   "Carrier_44_SpareOutput(5_5)" AT %I2568.5 : Bool;   // SPARE OUTPUT
   "Carrier_44_SpareOutput(5_6)" AT %I2568.6 : Bool;   // SPARE OUTPUT
   "Carrier_44_SpareOutput(5_7)" AT %I2568.7 : Bool;   // SPARE OUTPUT
   "Carrier_44_ActualSpeed" AT %IW2570 : Word;   // ACTUAL SPEED
   "Carrier_44_CarrierDriveAlarm" AT %IW2572 : Word;   // CARRIER DRIVE ALARM
   "Carrier_44_CarrierDriveWarning" AT %IW2574 : Word;   // CARRIER DRIVE WARNING
   "Carrier_45_Status" AT %IW2600 : Word;   // CARRIER STATUS WORD
   "Carrier_45_Status.0" AT %I2600.0 : Bool;   // HEARTBEAT
   "Carrier_45_Status.1" AT %I2600.1 : Bool;   // MANUAL
   "Carrier_45_Status.2" AT %I2600.2 : Bool;   // IN_AUTO
   "Carrier_45_Status.3" AT %I2600.3 : Bool;   // POSITIONING_COMPLETE
   "Carrier_45_Status.4" AT %I2600.4 : Bool;   // PRODUCTION HOLD
   "Carrier_45_Status.5" AT %I2600.5 : Bool;   // CARRIER MOVING FORWARD
   "Carrier_45_Status.6" AT %I2600.6 : Bool;   // CARRIER MOVING REVERSE
   "Carrier_45_Status.7" AT %I2600.7 : Bool;   // CARRIER FAULT
   "Carrier_45_Status.8" AT %I2601.0 : Bool;   // CRASH DETECT TRIPPED
   "Carrier_45_Status.9" AT %I2601.1 : Bool;
   "Carrier_45_Status.10" AT %I2601.2 : Bool;
   "Carrier_45_Status.11" AT %I2601.3 : Bool;
   "Carrier_45_Status.12" AT %I2601.4 : Bool;
   "Carrier_45_Status.13" AT %I2601.5 : Bool;
   "Carrier_45_Status.14" AT %I2601.6 : Bool;
   "Carrier_45_Status.15" AT %I2601.7 : Bool;
   "Carrier_45_SDCFaultCode" AT %IW2602 : Word;   // SDC FAULT CODE
   "Carrier_45_CarrierPosition" AT %ID2604 : DWord;   // CARRIER POSITION
   "Carrier_45_CarrierNumber" AT %IW2608 : Word;   // CARRIER NUMBER
   "Carrier_45_G120DControlWord" AT %IW2610 : Word;   // G120D_STW1_CONTROL
   "Carrier_45_G120DControlWord.0" AT %I2610.0 : Bool;   // Bit_00_ON
   "Carrier_45_G120DControlWord.1" AT %I2610.1 : Bool;   // Bit_01_AUS2_INH
   "Carrier_45_G120DControlWord.2" AT %I2610.2 : Bool;   // Bit_02_AUS3_STOP
   "Carrier_45_G120DControlWord.3" AT %I2610.3 : Bool;   // Bit_03_EN
   "Carrier_45_G120DControlWord.4" AT %I2610.4 : Bool;   // Bit_04_EN_RAMP
   "Carrier_45_G120DControlWord.5" AT %I2610.5 : Bool;   // Bit_05_START_RAMP
   "Carrier_45_G120DControlWord.6" AT %I2610.6 : Bool;   // Bit_06_SETPOINT
   "Carrier_45_G120DControlWord.7" AT %I2610.7 : Bool;   // Bit_07_RESET
   "Carrier_45_G120DControlWord.8" AT %I2611.0 : Bool;   // Bit_08_JOG_R
   "Carrier_45_G120DControlWord.9" AT %I2611.1 : Bool;   // Bit_09_JOG_L
   "Carrier_45_G120DControlWord.10" AT %I2611.2 : Bool;   // Bit_10_CONTR_PLC
   "Carrier_45_G120DControlWord.11" AT %I2611.3 : Bool;   // Bit_11_REVERSE
   "Carrier_45_G120DControlWord.12" AT %I2611.4 : Bool;   // Bit_12_BRAKE_RELEASE
   "Carrier_45_G120DControlWord.13" AT %I2611.5 : Bool;   // Bit_13_DDS
   "Carrier_45_G120DControlWord.14" AT %I2611.6 : Bool;   // Bit_14_DO0
   "Carrier_45_G120DControlWord.15" AT %I2611.7 : Bool;   // Bit_15_DO1
   "Carrier_45_G120DStatusWord" AT %IW2612 : Word;   // G120D_ZSW1_STATUS
   "Carrier_45_G120DStatusWord.0" AT %I2612.0 : Bool;   // Bit_00_READY_RUN
   "Carrier_45_G120DStatusWord.1" AT %I2612.1 : Bool;   // Bit_01_READY_ON
   "Carrier_45_G120DStatusWord.2" AT %I2612.2 : Bool;   // Bit_02_ENABLE
   "Carrier_45_G120DStatusWord.3" AT %I2612.3 : Bool;   // Bit_03_FAULT
   "Carrier_45_G120DStatusWord.4" AT %I2612.4 : Bool;   // Bit_04_OFF2
   "Carrier_45_G120DStatusWord.5" AT %I2612.5 : Bool;   // Bit_05_OFF3
   "Carrier_45_G120DStatusWord.6" AT %I2612.6 : Bool;   // Bit_06_LOCK_OUT
   "Carrier_45_G120DStatusWord.7" AT %I2612.7 : Bool;   // Bit_07_WARN
   "Carrier_45_G120DStatusWord.8" AT %I2613.0 : Bool;   // Bit_08_NO_DEVIATION
   "Carrier_45_G120DStatusWord.9" AT %I2613.1 : Bool;   // Bit_09_CONTR_PLC
   "Carrier_45_G120DStatusWord.10" AT %I2613.2 : Bool;   // Bit_10_F_MAX
   "Carrier_45_G120DStatusWord.11" AT %I2613.3 : Bool;   // Bit_11_LIMIT_REACHED
   "Carrier_45_G120DStatusWord.12" AT %I2613.4 : Bool;   // Bit_12_BRAKE_OPEN
   "Carrier_45_G120DStatusWord.13" AT %I2613.5 : Bool;   // Bit_13_NO_OVERTEMP
   "Carrier_45_G120DStatusWord.14" AT %I2613.6 : Bool;   // Bit_14_CW_CCW
   "Carrier_45_G120DStatusWord.15" AT %I2613.7 : Bool;   // Bit_15_OVERL
   "Carrier_45_Slot2_Input" AT %IW2614 : Word;   // SLOT 2 INPUT WORD
   "Carrier_45_CrashDetectSW" AT %I2614.0 : Bool;   // CRASH DETECT SW
   "Carrier_45_SpareSafetyInput(2_1)" AT %I2614.1 : Bool;   // SPARE SAFETY INPUT
   "Carrier_45_SpareSafetyInput(2_2)" AT %I2614.2 : Bool;   // SPARE SAFETY INPUT
   "Carrier_45_SpareSafetyInput(2_3)" AT %I2614.3 : Bool;   // SPARE SAFETY INPUT
   "Carrier_45_SpareSafetyInput(2_4)" AT %I2614.4 : Bool;   // SPARE SAFETY INPUT
   "Carrier_45_SpareSafetyInput(2_5)" AT %I2614.5 : Bool;   // SPARE SAFETY INPUT
   "Carrier_45_SpareSafetyInput(2_6)" AT %I2614.6 : Bool;   // SPARE SAFETY INPUT
   "Carrier_45_SpareSafetyInput(2_7)" AT %I2614.7 : Bool;   // SPARE SAFETY INPUT
   "Carrier_45_Slot3_SafetyOutput" AT %IW2615 : Word;   // SLOT 3 SAFETY OUTPUT WORD
   "Carrier_45_Crash_Detect_OK" AT %I2615.0 : Bool;   // CARRIER CRASH DETECT
   "Carrier_45_SpareSafetyOutput(3_1)" AT %I2615.1 : Bool;   // SPARE SAFETY OUTPUT
   "Carrier_45_SpareSafetyOutput(3_2)" AT %I2615.2 : Bool;   // SPARE SAFETY OUTPUT
   "Carrier_45_SpareSafetyOutput(3_3)" AT %I2615.3 : Bool;   // SPARE SAFETY OUTPUT
   "Carrier_45_SpareSafetyOutput(3_4)" AT %I2615.4 : Bool;   // SPARE SAFETY OUTPUT
   "Carrier_45_SpareSafetyOutput(3_5)" AT %I2615.5 : Bool;   // SPARE SAFETY OUTPUT
   "Carrier_45_SpareSafetyOutput(3_6)" AT %I2615.6 : Bool;   // SPARE SAFETY OUTPUT
   "Carrier_45_SpareSafetyOutput(3_7)" AT %I2615.7 : Bool;   // SPARE SAFETY OUTPUT
   "Carrier_45_Slot4_Input" AT %IW2616 : Word;   // SLOT 4 INPUT WORD
   "Carrier_45_480VPowerOn_MDCB1" AT %I2616.0 : Bool;   // 480 VAC POWER ON MDCB 1
   "Carrier_45_SpareInput(4_1)" AT %I2616.1 : Bool;   // SPARE INPUT
   "Carrier_45_SpareInput(4_2)" AT %I2616.2 : Bool;   // SPARE INPUT
   "Carrier_45_SitopSelectStatus" AT %I2616.3 : Bool;   // SITOP SELECT STATUS
   "Carrier_45_DCsupplyOnPSCB2" AT %I2616.4 : Bool;   // DC SUPPLY ON PSCB 2
   "Carrier_45_SpareInput(4_5)" AT %I2616.5 : Bool;   // SPARE INPUT
   "Carrier_45_SpareInput(4_6)" AT %I2616.6 : Bool;   // SPARE INPUT
   "Carrier_45_SpareInput(4_7)" AT %I2616.7 : Bool;   // SPARE INPUT
   "Carrier_45_PB1_ProdHoldLH" AT %I2617.0 : Bool;   // PB 1 PRODUCTION HOLD LH
   "Carrier_45_PB2_ResetLH" AT %I2617.1 : Bool;   // PB 2 RESET LH
   "Carrier_45_PB3_ProdHoldRH" AT %I2617.2 : Bool;   // PB 3 PRODUCTION HOLD RH
   "Carrier_45_PB4_ResetRH" AT %I2617.3 : Bool;   // PB 4 RESET RH
   "Carrier_45_SpareInput(4_14)" AT %I2617.4 : Bool;   // SPARE INPUT
   "Carrier_45_SpareInput(4_15)" AT %I2617.5 : Bool;   // SPARE INPUT
   "Carrier_45_SpareInput(4_16)" AT %I2617.6 : Bool;   // SPARE INPUT
   "Carrier_45_SpareInput(4_17)" AT %I2617.7 : Bool;   // SPARE INPUT
   "Carrier_45_Slot5_Output" AT %IW2618 : Word;   // SLOT 5 OUTPUT WORD
   "Carrier_45_IRD400_HMI_24VDC_ENABLE" AT %I2618.0 : Bool;   // IRD 400 PANEL HMI 24V DC POWER
   "Carrier_45_FaultLight_LH" AT %I2618.1 : Bool;   // FAULT LIGHT LH
   "Carrier_45_RunLight_LH" AT %I2618.2 : Bool;   // RUN LIGHT LH
   "Carrier_45_FaultLight_RH" AT %I2618.3 : Bool;   // FAULT LIGHT RH
   "Carrier_45_RunLight_RH" AT %I2618.4 : Bool;   // RUN LIGHT RH
   "Carrier_45_SpareOutput(5_5)" AT %I2618.5 : Bool;   // SPARE OUTPUT
   "Carrier_45_SpareOutput(5_6)" AT %I2618.6 : Bool;   // SPARE OUTPUT
   "Carrier_45_SpareOutput(5_7)" AT %I2618.7 : Bool;   // SPARE OUTPUT
   "Carrier_45_ActualSpeed" AT %IW2620 : Word;   // ACTUAL SPEED
   "Carrier_45_CarrierDriveAlarm" AT %IW2622 : Word;   // CARRIER DRIVE ALARM
   "Carrier_45_CarrierDriveWarning" AT %IW2624 : Word;   // CARRIER DRIVE WARNING
   "Carrier_46_Status" AT %IW2650 : Word;   // CARRIER STATUS WORD
   "Carrier_46_Status.0" AT %I2650.0 : Bool;   // HEARTBEAT
   "Carrier_46_Status.1" AT %I2650.1 : Bool;   // MANUAL
   "Carrier_46_Status.2" AT %I2650.2 : Bool;   // IN_AUTO
   "Carrier_46_Status.3" AT %I2650.3 : Bool;   // POSITIONING_COMPLETE
   "Carrier_46_Status.4" AT %I2650.4 : Bool;   // PRODUCTION HOLD
   "Carrier_46_Status.5" AT %I2650.5 : Bool;   // CARRIER MOVING FORWARD
   "Carrier_46_Status.6" AT %I2650.6 : Bool;   // CARRIER MOVING REVERSE
   "Carrier_46_Status.7" AT %I2650.7 : Bool;   // CARRIER FAULT
   "Carrier_46_Status.8" AT %I2651.0 : Bool;   // CRASH DETECT TRIPPED
   "Carrier_46_Status.9" AT %I2651.1 : Bool;
   "Carrier_46_Status.10" AT %I2651.2 : Bool;
   "Carrier_46_Status.11" AT %I2651.3 : Bool;
   "Carrier_46_Status.12" AT %I2651.4 : Bool;
   "Carrier_46_Status.13" AT %I2651.5 : Bool;
   "Carrier_46_Status.14" AT %I2651.6 : Bool;
   "Carrier_46_Status.15" AT %I2651.7 : Bool;
   "Carrier_46_SDCFaultCode" AT %IW2652 : Word;   // SDC FAULT CODE
   "Carrier_46_CarrierPosition" AT %ID2654 : DWord;   // CARRIER POSITION
   "Carrier_46_CarrierNumber" AT %IW2658 : Word;   // CARRIER NUMBER
   "Carrier_46_G120DControlWord" AT %IW2660 : Word;   // G120D_STW1_CONTROL
   "Carrier_46_G120DControlWord.0" AT %I2660.0 : Bool;   // Bit_00_ON
   "Carrier_46_G120DControlWord.1" AT %I2660.1 : Bool;   // Bit_01_AUS2_INH
   "Carrier_46_G120DControlWord.2" AT %I2660.2 : Bool;   // Bit_02_AUS3_STOP
   "Carrier_46_G120DControlWord.3" AT %I2660.3 : Bool;   // Bit_03_EN
   "Carrier_46_G120DControlWord.4" AT %I2660.4 : Bool;   // Bit_04_EN_RAMP
   "Carrier_46_G120DControlWord.5" AT %I2660.5 : Bool;   // Bit_05_START_RAMP
   "Carrier_46_G120DControlWord.6" AT %I2660.6 : Bool;   // Bit_06_SETPOINT
   "Carrier_46_G120DControlWord.7" AT %I2660.7 : Bool;   // Bit_07_RESET
   "Carrier_46_G120DControlWord.8" AT %I2661.0 : Bool;   // Bit_08_JOG_R
   "Carrier_46_G120DControlWord.9" AT %I2661.1 : Bool;   // Bit_09_JOG_L
   "Carrier_46_G120DControlWord.10" AT %I2661.2 : Bool;   // Bit_10_CONTR_PLC
   "Carrier_46_G120DControlWord.11" AT %I2661.3 : Bool;   // Bit_11_REVERSE
   "Carrier_46_G120DControlWord.12" AT %I2661.4 : Bool;   // Bit_12_BRAKE_RELEASE
   "Carrier_46_G120DControlWord.13" AT %I2661.5 : Bool;   // Bit_13_DDS
   "Carrier_46_G120DControlWord.14" AT %I2661.6 : Bool;   // Bit_14_DO0
   "Carrier_46_G120DControlWord.15" AT %I2661.7 : Bool;   // Bit_15_DO1
   "Carrier_46_G120DStatusWord" AT %IW2662 : Word;   // G120D_ZSW1_STATUS
   "Carrier_46_G120DStatusWord.0" AT %I2662.0 : Bool;   // Bit_00_READY_RUN
   "Carrier_46_G120DStatusWord.1" AT %I2662.1 : Bool;   // Bit_01_READY_ON
   "Carrier_46_G120DStatusWord.2" AT %I2662.2 : Bool;   // Bit_02_ENABLE
   "Carrier_46_G120DStatusWord.3" AT %I2662.3 : Bool;   // Bit_03_FAULT
   "Carrier_46_G120DStatusWord.4" AT %I2662.4 : Bool;   // Bit_04_OFF2
   "Carrier_46_G120DStatusWord.5" AT %I2662.5 : Bool;   // Bit_05_OFF3
   "Carrier_46_G120DStatusWord.6" AT %I2662.6 : Bool;   // Bit_06_LOCK_OUT
   "Carrier_46_G120DStatusWord.7" AT %I2662.7 : Bool;   // Bit_07_WARN
   "Carrier_46_G120DStatusWord.8" AT %I2663.0 : Bool;   // Bit_08_NO_DEVIATION
   "Carrier_46_G120DStatusWord.9" AT %I2663.1 : Bool;   // Bit_09_CONTR_PLC
   "Carrier_46_G120DStatusWord.10" AT %I2663.2 : Bool;   // Bit_10_F_MAX
   "Carrier_46_G120DStatusWord.11" AT %I2663.3 : Bool;   // Bit_11_LIMIT_REACHED
   "Carrier_46_G120DStatusWord.12" AT %I2663.4 : Bool;   // Bit_12_BRAKE_OPEN
   "Carrier_46_G120DStatusWord.13" AT %I2663.5 : Bool;   // Bit_13_NO_OVERTEMP
   "Carrier_46_G120DStatusWord.14" AT %I2663.6 : Bool;   // Bit_14_CW_CCW
   "Carrier_46_G120DStatusWord.15" AT %I2663.7 : Bool;   // Bit_15_OVERL
   "Carrier_46_Slot2_Input" AT %IW2664 : Word;   // SLOT 2 INPUT WORD
   "Carrier_46_CrashDetectSW" AT %I2664.0 : Bool;   // CRASH DETECT SW
   "Carrier_46_SpareSafetyInput(2_1)" AT %I2664.1 : Bool;   // SPARE SAFETY INPUT
   "Carrier_46_SpareSafetyInput(2_2)" AT %I2664.2 : Bool;   // SPARE SAFETY INPUT
   "Carrier_46_SpareSafetyInput(2_3)" AT %I2664.3 : Bool;   // SPARE SAFETY INPUT
   "Carrier_46_SpareSafetyInput(2_4)" AT %I2664.4 : Bool;   // SPARE SAFETY INPUT
   "Carrier_46_SpareSafetyInput(2_5)" AT %I2664.5 : Bool;   // SPARE SAFETY INPUT
   "Carrier_46_SpareSafetyInput(2_6)" AT %I2664.6 : Bool;   // SPARE SAFETY INPUT
   "Carrier_46_SpareSafetyInput(2_7)" AT %I2664.7 : Bool;   // SPARE SAFETY INPUT
   "Carrier_46_Slot3_SafetyOutput" AT %IW2665 : Word;   // SLOT 3 SAFETY OUTPUT WORD
   "Carrier_46_Crash_Detect_OK" AT %I2665.0 : Bool;   // CARRIER CRASH DETECT
   "Carrier_46_SpareSafetyOutput(3_1)" AT %I2665.1 : Bool;   // SPARE SAFETY OUTPUT
   "Carrier_46_SpareSafetyOutput(3_2)" AT %I2665.2 : Bool;   // SPARE SAFETY OUTPUT
   "Carrier_46_SpareSafetyOutput(3_3)" AT %I2665.3 : Bool;   // SPARE SAFETY OUTPUT
   "Carrier_46_SpareSafetyOutput(3_4)" AT %I2665.4 : Bool;   // SPARE SAFETY OUTPUT
   "Carrier_46_SpareSafetyOutput(3_5)" AT %I2665.5 : Bool;   // SPARE SAFETY OUTPUT
   "Carrier_46_SpareSafetyOutput(3_6)" AT %I2665.6 : Bool;   // SPARE SAFETY OUTPUT
   "Carrier_46_SpareSafetyOutput(3_7)" AT %I2665.7 : Bool;   // SPARE SAFETY OUTPUT
   "Carrier_46_Slot4_Input" AT %IW2666 : Word;   // SLOT 4 INPUT WORD
   "Carrier_46_480VPowerOn_MDCB1" AT %I2666.0 : Bool;   // 480 VAC POWER ON MDCB 1
   "Carrier_46_SpareInput(4_1)" AT %I2666.1 : Bool;   // SPARE INPUT
   "Carrier_46_SpareInput(4_2)" AT %I2666.2 : Bool;   // SPARE INPUT
   "Carrier_46_SitopSelectStatus" AT %I2666.3 : Bool;   // SITOP SELECT STATUS
   "Carrier_46_DCsupplyOnPSCB2" AT %I2666.4 : Bool;   // DC SUPPLY ON PSCB 2
   "Carrier_46_SpareInput(4_5)" AT %I2666.5 : Bool;   // SPARE INPUT
   "Carrier_46_SpareInput(4_6)" AT %I2666.6 : Bool;   // SPARE INPUT
   "Carrier_46_SpareInput(4_7)" AT %I2666.7 : Bool;   // SPARE INPUT
   "Carrier_46_PB1_ProdHoldLH" AT %I2667.0 : Bool;   // PB 1 PRODUCTION HOLD LH
   "Carrier_46_PB2_ResetLH" AT %I2667.1 : Bool;   // PB 2 RESET LH
   "Carrier_46_PB3_ProdHoldRH" AT %I2667.2 : Bool;   // PB 3 PRODUCTION HOLD RH
   "Carrier_46_PB4_ResetRH" AT %I2667.3 : Bool;   // PB 4 RESET RH
   "Carrier_46_SpareInput(4_14)" AT %I2667.4 : Bool;   // SPARE INPUT
   "Carrier_46_SpareInput(4_15)" AT %I2667.5 : Bool;   // SPARE INPUT
   "Carrier_46_SpareInput(4_16)" AT %I2667.6 : Bool;   // SPARE INPUT
   "Carrier_46_SpareInput(4_17)" AT %I2667.7 : Bool;   // SPARE INPUT
   "Carrier_46_Slot5_Output" AT %IW2668 : Word;   // SLOT 5 OUTPUT WORD
   "Carrier_46_IRD400_HMI_24VDC_ENABLE" AT %I2668.0 : Bool;   // IRD 400 PANEL HMI 24V DC POWER
   "Carrier_46_FaultLight_LH" AT %I2668.1 : Bool;   // FAULT LIGHT LH
   "Carrier_46_RunLight_LH" AT %I2668.2 : Bool;   // RUN LIGHT LH
   "Carrier_46_FaultLight_RH" AT %I2668.3 : Bool;   // FAULT LIGHT RH
   "Carrier_46_RunLight_RH" AT %I2668.4 : Bool;   // RUN LIGHT RH
   "Carrier_46_SpareOutput(5_5)" AT %I2668.5 : Bool;   // SPARE OUTPUT
   "Carrier_46_SpareOutput(5_6)" AT %I2668.6 : Bool;   // SPARE OUTPUT
   "Carrier_46_SpareOutput(5_7)" AT %I2668.7 : Bool;   // SPARE OUTPUT
   "Carrier_46_ActualSpeed" AT %IW2670 : Word;   // ACTUAL SPEED
   "Carrier_46_CarrierDriveAlarm" AT %IW2672 : Word;   // CARRIER DRIVE ALARM
   "Carrier_46_CarrierDriveWarning" AT %IW2674 : Word;   // CARRIER DRIVE WARNING
   "Carrier_47_Status" AT %IW2700 : Word;   // CARRIER STATUS WORD
   "Carrier_47_Status.0" AT %I2700.0 : Bool;   // HEARTBEAT
   "Carrier_47_Status.1" AT %I2700.1 : Bool;   // MANUAL
   "Carrier_47_Status.2" AT %I2700.2 : Bool;   // IN_AUTO
   "Carrier_47_Status.3" AT %I2700.3 : Bool;   // POSITIONING_COMPLETE
   "Carrier_47_Status.4" AT %I2700.4 : Bool;   // PRODUCTION HOLD
   "Carrier_47_Status.5" AT %I2700.5 : Bool;   // CARRIER MOVING FORWARD
   "Carrier_47_Status.6" AT %I2700.6 : Bool;   // CARRIER MOVING REVERSE
   "Carrier_47_Status.7" AT %I2700.7 : Bool;   // CARRIER FAULT
   "Carrier_47_Status.8" AT %I2701.0 : Bool;   // CRASH DETECT TRIPPED
   "Carrier_47_Status.9" AT %I2701.1 : Bool;
   "Carrier_47_Status.10" AT %I2701.2 : Bool;
   "Carrier_47_Status.11" AT %I2701.3 : Bool;
   "Carrier_47_Status.12" AT %I2701.4 : Bool;
   "Carrier_47_Status.13" AT %I2701.5 : Bool;
   "Carrier_47_Status.14" AT %I2701.6 : Bool;
   "Carrier_47_Status.15" AT %I2701.7 : Bool;
   "Carrier_47_SDCFaultCode" AT %IW2702 : Word;   // SDC FAULT CODE
   "Carrier_47_CarrierPosition" AT %ID2704 : DWord;   // CARRIER POSITION
   "Carrier_47_CarrierNumber" AT %IW2708 : Word;   // CARRIER NUMBER
   "Carrier_47_G120DControlWord" AT %IW2710 : Word;   // G120D_STW1_CONTROL
   "Carrier_47_G120DControlWord.0" AT %I2710.0 : Bool;   // Bit_00_ON
   "Carrier_47_G120DControlWord.1" AT %I2710.1 : Bool;   // Bit_01_AUS2_INH
   "Carrier_47_G120DControlWord.2" AT %I2710.2 : Bool;   // Bit_02_AUS3_STOP
   "Carrier_47_G120DControlWord.3" AT %I2710.3 : Bool;   // Bit_03_EN
   "Carrier_47_G120DControlWord.4" AT %I2710.4 : Bool;   // Bit_04_EN_RAMP
   "Carrier_47_G120DControlWord.5" AT %I2710.5 : Bool;   // Bit_05_START_RAMP
   "Carrier_47_G120DControlWord.6" AT %I2710.6 : Bool;   // Bit_06_SETPOINT
   "Carrier_47_G120DControlWord.7" AT %I2710.7 : Bool;   // Bit_07_RESET
   "Carrier_47_G120DControlWord.8" AT %I2711.0 : Bool;   // Bit_08_JOG_R
   "Carrier_47_G120DControlWord.9" AT %I2711.1 : Bool;   // Bit_09_JOG_L
   "Carrier_47_G120DControlWord.10" AT %I2711.2 : Bool;   // Bit_10_CONTR_PLC
   "Carrier_47_G120DControlWord.11" AT %I2711.3 : Bool;   // Bit_11_REVERSE
   "Carrier_47_G120DControlWord.12" AT %I2711.4 : Bool;   // Bit_12_BRAKE_RELEASE
   "Carrier_47_G120DControlWord.13" AT %I2711.5 : Bool;   // Bit_13_DDS
   "Carrier_47_G120DControlWord.14" AT %I2711.6 : Bool;   // Bit_14_DO0
   "Carrier_47_G120DControlWord.15" AT %I2711.7 : Bool;   // Bit_15_DO1
   "Carrier_47_G120DStatusWord" AT %IW2712 : Word;   // G120D_ZSW1_STATUS
   "Carrier_47_G120DStatusWord.0" AT %I2712.0 : Bool;   // Bit_00_READY_RUN
   "Carrier_47_G120DStatusWord.1" AT %I2712.1 : Bool;   // Bit_01_READY_ON
   "Carrier_47_G120DStatusWord.2" AT %I2712.2 : Bool;   // Bit_02_ENABLE
   "Carrier_47_G120DStatusWord.3" AT %I2712.3 : Bool;   // Bit_03_FAULT
   "Carrier_47_G120DStatusWord.4" AT %I2712.4 : Bool;   // Bit_04_OFF2
   "Carrier_47_G120DStatusWord.5" AT %I2712.5 : Bool;   // Bit_05_OFF3
   "Carrier_47_G120DStatusWord.6" AT %I2712.6 : Bool;   // Bit_06_LOCK_OUT
   "Carrier_47_G120DStatusWord.7" AT %I2712.7 : Bool;   // Bit_07_WARN
   "Carrier_47_G120DStatusWord.8" AT %I2713.0 : Bool;   // Bit_08_NO_DEVIATION
   "Carrier_47_G120DStatusWord.9" AT %I2713.1 : Bool;   // Bit_09_CONTR_PLC
   "Carrier_47_G120DStatusWord.10" AT %I2713.2 : Bool;   // Bit_10_F_MAX
   "Carrier_47_G120DStatusWord.11" AT %I2713.3 : Bool;   // Bit_11_LIMIT_REACHED
   "Carrier_47_G120DStatusWord.12" AT %I2713.4 : Bool;   // Bit_12_BRAKE_OPEN
   "Carrier_47_G120DStatusWord.13" AT %I2713.5 : Bool;   // Bit_13_NO_OVERTEMP
   "Carrier_47_G120DStatusWord.14" AT %I2713.6 : Bool;   // Bit_14_CW_CCW
   "Carrier_47_G120DStatusWord.15" AT %I2713.7 : Bool;   // Bit_15_OVERL
   "Carrier_47_Slot2_Input" AT %IW2714 : Word;   // SLOT 2 INPUT WORD
   "Carrier_47_CrashDetectSW" AT %I2714.0 : Bool;   // CRASH DETECT SW
   "Carrier_47_SpareSafetyInput(2_1)" AT %I2714.1 : Bool;   // SPARE SAFETY INPUT
   "Carrier_47_SpareSafetyInput(2_2)" AT %I2714.2 : Bool;   // SPARE SAFETY INPUT
   "Carrier_47_SpareSafetyInput(2_3)" AT %I2714.3 : Bool;   // SPARE SAFETY INPUT
   "Carrier_47_SpareSafetyInput(2_4)" AT %I2714.4 : Bool;   // SPARE SAFETY INPUT
   "Carrier_47_SpareSafetyInput(2_5)" AT %I2714.5 : Bool;   // SPARE SAFETY INPUT
   "Carrier_47_SpareSafetyInput(2_6)" AT %I2714.6 : Bool;   // SPARE SAFETY INPUT
   "Carrier_47_SpareSafetyInput(2_7)" AT %I2714.7 : Bool;   // SPARE SAFETY INPUT
   "Carrier_47_Slot3_SafetyOutput" AT %IW2715 : Word;   // SLOT 3 SAFETY OUTPUT WORD
   "Carrier_47_Crash_Detect_OK" AT %I2715.0 : Bool;   // CARRIER CRASH DETECT
   "Carrier_47_SpareSafetyOutput(3_1)" AT %I2715.1 : Bool;   // SPARE SAFETY OUTPUT
   "Carrier_47_SpareSafetyOutput(3_2)" AT %I2715.2 : Bool;   // SPARE SAFETY OUTPUT
   "Carrier_47_SpareSafetyOutput(3_3)" AT %I2715.3 : Bool;   // SPARE SAFETY OUTPUT
   "Carrier_47_SpareSafetyOutput(3_4)" AT %I2715.4 : Bool;   // SPARE SAFETY OUTPUT
   "Carrier_47_SpareSafetyOutput(3_5)" AT %I2715.5 : Bool;   // SPARE SAFETY OUTPUT
   "Carrier_47_SpareSafetyOutput(3_6)" AT %I2715.6 : Bool;   // SPARE SAFETY OUTPUT
   "Carrier_47_SpareSafetyOutput(3_7)" AT %I2715.7 : Bool;   // SPARE SAFETY OUTPUT
   "Carrier_47_Slot4_Input" AT %IW2716 : Word;   // SLOT 4 INPUT WORD
   "Carrier_47_480VPowerOn_MDCB1" AT %I2716.0 : Bool;   // 480 VAC POWER ON MDCB 1
   "Carrier_47_SpareInput(4_1)" AT %I2716.1 : Bool;   // SPARE INPUT
   "Carrier_47_SpareInput(4_2)" AT %I2716.2 : Bool;   // SPARE INPUT
   "Carrier_47_SitopSelectStatus" AT %I2716.3 : Bool;   // SITOP SELECT STATUS
   "Carrier_47_DCsupplyOnPSCB2" AT %I2716.4 : Bool;   // DC SUPPLY ON PSCB 2
   "Carrier_47_SpareInput(4_5)" AT %I2716.5 : Bool;   // SPARE INPUT
   "Carrier_47_SpareInput(4_6)" AT %I2716.6 : Bool;   // SPARE INPUT
   "Carrier_47_SpareInput(4_7)" AT %I2716.7 : Bool;   // SPARE INPUT
   "Carrier_47_PB1_ProdHoldLH" AT %I2717.0 : Bool;   // PB 1 PRODUCTION HOLD LH
   "Carrier_47_PB2_ResetLH" AT %I2717.1 : Bool;   // PB 2 RESET LH
   "Carrier_47_PB3_ProdHoldRH" AT %I2717.2 : Bool;   // PB 3 PRODUCTION HOLD RH
   "Carrier_47_PB4_ResetRH" AT %I2717.3 : Bool;   // PB 4 RESET RH
   "Carrier_47_SpareInput(4_14)" AT %I2717.4 : Bool;   // SPARE INPUT
   "Carrier_47_SpareInput(4_15)" AT %I2717.5 : Bool;   // SPARE INPUT
   "Carrier_47_SpareInput(4_16)" AT %I2717.6 : Bool;   // SPARE INPUT
   "Carrier_47_SpareInput(4_17)" AT %I2717.7 : Bool;   // SPARE INPUT
   "Carrier_47_Slot5_Output" AT %IW2718 : Word;   // SLOT 5 OUTPUT WORD
   "Carrier_47_IRD400_HMI_24VDC_ENABLE" AT %I2718.0 : Bool;   // IRD 400 PANEL HMI 24V DC POWER
   "Carrier_47_FaultLight_LH" AT %I2718.1 : Bool;   // FAULT LIGHT LH
   "Carrier_47_RunLight_LH" AT %I2718.2 : Bool;   // RUN LIGHT LH
   "Carrier_47_FaultLight_RH" AT %I2718.3 : Bool;   // FAULT LIGHT RH
   "Carrier_47_RunLight_RH" AT %I2718.4 : Bool;   // RUN LIGHT RH
   "Carrier_47_SpareOutput(5_5)" AT %I2718.5 : Bool;   // SPARE OUTPUT
   "Carrier_47_SpareOutput(5_6)" AT %I2718.6 : Bool;   // SPARE OUTPUT
   "Carrier_47_SpareOutput(5_7)" AT %I2718.7 : Bool;   // SPARE OUTPUT
   "Carrier_47_ActualSpeed" AT %IW2720 : Word;   // ACTUAL SPEED
   "Carrier_47_CarrierDriveAlarm" AT %IW2722 : Word;   // CARRIER DRIVE ALARM
   "Carrier_47_CarrierDriveWarning" AT %IW2724 : Word;   // CARRIER DRIVE WARNING
   "Carrier_48_Status" AT %IW2750 : Word;   // CARRIER STATUS WORD
   "Carrier_48_Status.0" AT %I2750.0 : Bool;   // HEARTBEAT
   "Carrier_48_Status.1" AT %I2750.1 : Bool;   // MANUAL
   "Carrier_48_Status.2" AT %I2750.2 : Bool;   // IN_AUTO
   "Carrier_48_Status.3" AT %I2750.3 : Bool;   // POSITIONING_COMPLETE
   "Carrier_48_Status.4" AT %I2750.4 : Bool;   // PRODUCTION HOLD
   "Carrier_48_Status.5" AT %I2750.5 : Bool;   // CARRIER MOVING FORWARD
   "Carrier_48_Status.6" AT %I2750.6 : Bool;   // CARRIER MOVING REVERSE
   "Carrier_48_Status.7" AT %I2750.7 : Bool;   // CARRIER FAULT
   "Carrier_48_Status.8" AT %I2751.0 : Bool;   // CRASH DETECT TRIPPED
   "Carrier_48_Status.9" AT %I2751.1 : Bool;
   "Carrier_48_Status.10" AT %I2751.2 : Bool;
   "Carrier_48_Status.11" AT %I2751.3 : Bool;
   "Carrier_48_Status.12" AT %I2751.4 : Bool;
   "Carrier_48_Status.13" AT %I2751.5 : Bool;
   "Carrier_48_Status.14" AT %I2751.6 : Bool;
   "Carrier_48_Status.15" AT %I2751.7 : Bool;
   "Carrier_48_SDCFaultCode" AT %IW2752 : Word;   // SDC FAULT CODE
   "Carrier_48_CarrierPosition" AT %ID2754 : DWord;   // CARRIER POSITION
   "Carrier_48_CarrierNumber" AT %IW2758 : Word;   // CARRIER NUMBER
   "Carrier_48_G120DControlWord" AT %IW2760 : Word;   // G120D_STW1_CONTROL
   "Carrier_48_G120DControlWord.0" AT %I2760.0 : Bool;   // Bit_00_ON
   "Carrier_48_G120DControlWord.1" AT %I2760.1 : Bool;   // Bit_01_AUS2_INH
   "Carrier_48_G120DControlWord.2" AT %I2760.2 : Bool;   // Bit_02_AUS3_STOP
   "Carrier_48_G120DControlWord.3" AT %I2760.3 : Bool;   // Bit_03_EN
   "Carrier_48_G120DControlWord.4" AT %I2760.4 : Bool;   // Bit_04_EN_RAMP
   "Carrier_48_G120DControlWord.5" AT %I2760.5 : Bool;   // Bit_05_START_RAMP
   "Carrier_48_G120DControlWord.6" AT %I2760.6 : Bool;   // Bit_06_SETPOINT
   "Carrier_48_G120DControlWord.7" AT %I2760.7 : Bool;   // Bit_07_RESET
   "Carrier_48_G120DControlWord.8" AT %I2761.0 : Bool;   // Bit_08_JOG_R
   "Carrier_48_G120DControlWord.9" AT %I2761.1 : Bool;   // Bit_09_JOG_L
   "Carrier_48_G120DControlWord.10" AT %I2761.2 : Bool;   // Bit_10_CONTR_PLC
   "Carrier_48_G120DControlWord.11" AT %I2761.3 : Bool;   // Bit_11_REVERSE
   "Carrier_48_G120DControlWord.12" AT %I2761.4 : Bool;   // Bit_12_BRAKE_RELEASE
   "Carrier_48_G120DControlWord.13" AT %I2761.5 : Bool;   // Bit_13_DDS
   "Carrier_48_G120DControlWord.14" AT %I2761.6 : Bool;   // Bit_14_DO0
   "Carrier_48_G120DControlWord.15" AT %I2761.7 : Bool;   // Bit_15_DO1
   "Carrier_48_G120DStatusWord" AT %IW2762 : Word;   // G120D_ZSW1_STATUS
   "Carrier_48_G120DStatusWord.0" AT %I2762.0 : Bool;   // Bit_00_READY_RUN
   "Carrier_48_G120DStatusWord.1" AT %I2762.1 : Bool;   // Bit_01_READY_ON
   "Carrier_48_G120DStatusWord.2" AT %I2762.2 : Bool;   // Bit_02_ENABLE
   "Carrier_48_G120DStatusWord.3" AT %I2762.3 : Bool;   // Bit_03_FAULT
   "Carrier_48_G120DStatusWord.4" AT %I2762.4 : Bool;   // Bit_04_OFF2
   "Carrier_48_G120DStatusWord.5" AT %I2762.5 : Bool;   // Bit_05_OFF3
   "Carrier_48_G120DStatusWord.6" AT %I2762.6 : Bool;   // Bit_06_LOCK_OUT
   "Carrier_48_G120DStatusWord.7" AT %I2762.7 : Bool;   // Bit_07_WARN
   "Carrier_48_G120DStatusWord.8" AT %I2763.0 : Bool;   // Bit_08_NO_DEVIATION
   "Carrier_48_G120DStatusWord.9" AT %I2763.1 : Bool;   // Bit_09_CONTR_PLC
   "Carrier_48_G120DStatusWord.10" AT %I2763.2 : Bool;   // Bit_10_F_MAX
   "Carrier_48_G120DStatusWord.11" AT %I2763.3 : Bool;   // Bit_11_LIMIT_REACHED
   "Carrier_48_G120DStatusWord.12" AT %I2763.4 : Bool;   // Bit_12_BRAKE_OPEN
   "Carrier_48_G120DStatusWord.13" AT %I2763.5 : Bool;   // Bit_13_NO_OVERTEMP
   "Carrier_48_G120DStatusWord.14" AT %I2763.6 : Bool;   // Bit_14_CW_CCW
   "Carrier_48_G120DStatusWord.15" AT %I2763.7 : Bool;   // Bit_15_OVERL
   "Carrier_48_Slot2_Input" AT %IW2764 : Word;   // SLOT 2 INPUT WORD
   "Carrier_48_CrashDetectSW" AT %I2764.0 : Bool;   // CRASH DETECT SW
   "Carrier_48_SpareSafetyInput(2_1)" AT %I2764.1 : Bool;   // SPARE SAFETY INPUT
   "Carrier_48_SpareSafetyInput(2_2)" AT %I2764.2 : Bool;   // SPARE SAFETY INPUT
   "Carrier_48_SpareSafetyInput(2_3)" AT %I2764.3 : Bool;   // SPARE SAFETY INPUT
   "Carrier_48_SpareSafetyInput(2_4)" AT %I2764.4 : Bool;   // SPARE SAFETY INPUT
   "Carrier_48_SpareSafetyInput(2_5)" AT %I2764.5 : Bool;   // SPARE SAFETY INPUT
   "Carrier_48_SpareSafetyInput(2_6)" AT %I2764.6 : Bool;   // SPARE SAFETY INPUT
   "Carrier_48_SpareSafetyInput(2_7)" AT %I2764.7 : Bool;   // SPARE SAFETY INPUT
   "Carrier_48_Slot3_SafetyOutput" AT %IW2765 : Word;   // SLOT 3 SAFETY OUTPUT WORD
   "Carrier_48_Crash_Detect_OK" AT %I2765.0 : Bool;   // CARRIER CRASH DETECT
   "Carrier_48_SpareSafetyOutput(3_1)" AT %I2765.1 : Bool;   // SPARE SAFETY OUTPUT
   "Carrier_48_SpareSafetyOutput(3_2)" AT %I2765.2 : Bool;   // SPARE SAFETY OUTPUT
   "Carrier_48_SpareSafetyOutput(3_3)" AT %I2765.3 : Bool;   // SPARE SAFETY OUTPUT
   "Carrier_48_SpareSafetyOutput(3_4)" AT %I2765.4 : Bool;   // SPARE SAFETY OUTPUT
   "Carrier_48_SpareSafetyOutput(3_5)" AT %I2765.5 : Bool;   // SPARE SAFETY OUTPUT
   "Carrier_48_SpareSafetyOutput(3_6)" AT %I2765.6 : Bool;   // SPARE SAFETY OUTPUT
   "Carrier_48_SpareSafetyOutput(3_7)" AT %I2765.7 : Bool;   // SPARE SAFETY OUTPUT
   "Carrier_48_Slot4_Input" AT %IW2766 : Word;   // SLOT 4 INPUT WORD
   "Carrier_48_480VPowerOn_MDCB1" AT %I2766.0 : Bool;   // 480 VAC POWER ON MDCB 1
   "Carrier_48_SpareInput(4_1)" AT %I2766.1 : Bool;   // SPARE INPUT
   "Carrier_48_SpareInput(4_2)" AT %I2766.2 : Bool;   // SPARE INPUT
   "Carrier_48_SitopSelectStatus" AT %I2766.3 : Bool;   // SITOP SELECT STATUS
   "Carrier_48_DCsupplyOnPSCB2" AT %I2766.4 : Bool;   // DC SUPPLY ON PSCB 2
   "Carrier_48_SpareInput(4_5)" AT %I2766.5 : Bool;   // SPARE INPUT
   "Carrier_48_SpareInput(4_6)" AT %I2766.6 : Bool;   // SPARE INPUT
   "Carrier_48_SpareInput(4_7)" AT %I2766.7 : Bool;   // SPARE INPUT
   "Carrier_48_PB1_ProdHoldLH" AT %I2767.0 : Bool;   // PB 1 PRODUCTION HOLD LH
   "Carrier_48_PB2_ResetLH" AT %I2767.1 : Bool;   // PB 2 RESET LH
   "Carrier_48_PB3_ProdHoldRH" AT %I2767.2 : Bool;   // PB 3 PRODUCTION HOLD RH
   "Carrier_48_PB4_ResetRH" AT %I2767.3 : Bool;   // PB 4 RESET RH
   "Carrier_48_SpareInput(4_14)" AT %I2767.4 : Bool;   // SPARE INPUT
   "Carrier_48_SpareInput(4_15)" AT %I2767.5 : Bool;   // SPARE INPUT
   "Carrier_48_SpareInput(4_16)" AT %I2767.6 : Bool;   // SPARE INPUT
   "Carrier_48_SpareInput(4_17)" AT %I2767.7 : Bool;   // SPARE INPUT
   "Carrier_48_Slot5_Output" AT %IW2768 : Word;   // SLOT 5 OUTPUT WORD
   "Carrier_48_IRD400_HMI_24VDC_ENABLE" AT %I2768.0 : Bool;   // IRD 400 PANEL HMI 24V DC POWER
   "Carrier_48_FaultLight_LH" AT %I2768.1 : Bool;   // FAULT LIGHT LH
   "Carrier_48_RunLight_LH" AT %I2768.2 : Bool;   // RUN LIGHT LH
   "Carrier_48_FaultLight_RH" AT %I2768.3 : Bool;   // FAULT LIGHT RH
   "Carrier_48_RunLight_RH" AT %I2768.4 : Bool;   // RUN LIGHT RH
   "Carrier_48_SpareOutput(5_5)" AT %I2768.5 : Bool;   // SPARE OUTPUT
   "Carrier_48_SpareOutput(5_6)" AT %I2768.6 : Bool;   // SPARE OUTPUT
   "Carrier_48_SpareOutput(5_7)" AT %I2768.7 : Bool;   // SPARE OUTPUT
   "Carrier_48_ActualSpeed" AT %IW2770 : Word;   // ACTUAL SPEED
   "Carrier_48_CarrierDriveAlarm" AT %IW2772 : Word;   // CARRIER DRIVE ALARM
   "Carrier_48_CarrierDriveWarning" AT %IW2774 : Word;   // CARRIER DRIVE WARNING
   "Carrier_49_Status" AT %IW2800 : Word;   // CARRIER STATUS WORD
   "Carrier_49_Status.0" AT %I2800.0 : Bool;   // HEARTBEAT
   "Carrier_49_Status.1" AT %I2800.1 : Bool;   // MANUAL
   "Carrier_49_Status.2" AT %I2800.2 : Bool;   // IN_AUTO
   "Carrier_49_Status.3" AT %I2800.3 : Bool;   // POSITIONING_COMPLETE
   "Carrier_49_Status.4" AT %I2800.4 : Bool;   // PRODUCTION HOLD
   "Carrier_49_Status.5" AT %I2800.5 : Bool;   // CARRIER MOVING FORWARD
   "Carrier_49_Status.6" AT %I2800.6 : Bool;   // CARRIER MOVING REVERSE
   "Carrier_49_Status.7" AT %I2800.7 : Bool;   // CARRIER FAULT
   "Carrier_49_Status.8" AT %I2801.0 : Bool;   // CRASH DETECT TRIPPED
   "Carrier_49_Status.9" AT %I2801.1 : Bool;
   "Carrier_49_Status.10" AT %I2801.2 : Bool;
   "Carrier_49_Status.11" AT %I2801.3 : Bool;
   "Carrier_49_Status.12" AT %I2801.4 : Bool;
   "Carrier_49_Status.13" AT %I2801.5 : Bool;
   "Carrier_49_Status.14" AT %I2801.6 : Bool;
   "Carrier_49_Status.15" AT %I2801.7 : Bool;
   "Carrier_49_SDCFaultCode" AT %IW2802 : Word;   // SDC FAULT CODE
   "Carrier_49_CarrierPosition" AT %ID2804 : DWord;   // CARRIER POSITION
   "Carrier_49_CarrierNumber" AT %IW2808 : Word;   // CARRIER NUMBER
   "Carrier_49_G120DControlWord" AT %IW2810 : Word;   // G120D_STW1_CONTROL
   "Carrier_49_G120DControlWord.0" AT %I2810.0 : Bool;   // Bit_00_ON
   "Carrier_49_G120DControlWord.1" AT %I2810.1 : Bool;   // Bit_01_AUS2_INH
   "Carrier_49_G120DControlWord.2" AT %I2810.2 : Bool;   // Bit_02_AUS3_STOP
   "Carrier_49_G120DControlWord.3" AT %I2810.3 : Bool;   // Bit_03_EN
   "Carrier_49_G120DControlWord.4" AT %I2810.4 : Bool;   // Bit_04_EN_RAMP
   "Carrier_49_G120DControlWord.5" AT %I2810.5 : Bool;   // Bit_05_START_RAMP
   "Carrier_49_G120DControlWord.6" AT %I2810.6 : Bool;   // Bit_06_SETPOINT
   "Carrier_49_G120DControlWord.7" AT %I2810.7 : Bool;   // Bit_07_RESET
   "Carrier_49_G120DControlWord.8" AT %I2811.0 : Bool;   // Bit_08_JOG_R
   "Carrier_49_G120DControlWord.9" AT %I2811.1 : Bool;   // Bit_09_JOG_L
   "Carrier_49_G120DControlWord.10" AT %I2811.2 : Bool;   // Bit_10_CONTR_PLC
   "Carrier_49_G120DControlWord.11" AT %I2811.3 : Bool;   // Bit_11_REVERSE
   "Carrier_49_G120DControlWord.12" AT %I2811.4 : Bool;   // Bit_12_BRAKE_RELEASE
   "Carrier_49_G120DControlWord.13" AT %I2811.5 : Bool;   // Bit_13_DDS
   "Carrier_49_G120DControlWord.14" AT %I2811.6 : Bool;   // Bit_14_DO0
   "Carrier_49_G120DControlWord.15" AT %I2811.7 : Bool;   // Bit_15_DO1
   "Carrier_49_G120DStatusWord" AT %IW2812 : Word;   // G120D_ZSW1_STATUS
   "Carrier_49_G120DStatusWord.0" AT %I2812.0 : Bool;   // Bit_00_READY_RUN
   "Carrier_49_G120DStatusWord.1" AT %I2812.1 : Bool;   // Bit_01_READY_ON
   "Carrier_49_G120DStatusWord.2" AT %I2812.2 : Bool;   // Bit_02_ENABLE
   "Carrier_49_G120DStatusWord.3" AT %I2812.3 : Bool;   // Bit_03_FAULT
   "Carrier_49_G120DStatusWord.4" AT %I2812.4 : Bool;   // Bit_04_OFF2
   "Carrier_49_G120DStatusWord.5" AT %I2812.5 : Bool;   // Bit_05_OFF3
   "Carrier_49_G120DStatusWord.6" AT %I2812.6 : Bool;   // Bit_06_LOCK_OUT
   "Carrier_49_G120DStatusWord.7" AT %I2812.7 : Bool;   // Bit_07_WARN
   "Carrier_49_G120DStatusWord.8" AT %I2813.0 : Bool;   // Bit_08_NO_DEVIATION
   "Carrier_49_G120DStatusWord.9" AT %I2813.1 : Bool;   // Bit_09_CONTR_PLC
   "Carrier_49_G120DStatusWord.10" AT %I2813.2 : Bool;   // Bit_10_F_MAX
   "Carrier_49_G120DStatusWord.11" AT %I2813.3 : Bool;   // Bit_11_LIMIT_REACHED
   "Carrier_49_G120DStatusWord.12" AT %I2813.4 : Bool;   // Bit_12_BRAKE_OPEN
   "Carrier_49_G120DStatusWord.13" AT %I2813.5 : Bool;   // Bit_13_NO_OVERTEMP
   "Carrier_49_G120DStatusWord.14" AT %I2813.6 : Bool;   // Bit_14_CW_CCW
   "Carrier_49_G120DStatusWord.15" AT %I2813.7 : Bool;   // Bit_15_OVERL